VERSION : 0.1
   VAR_INPUT
      OFF_SQ : Bool := false;   // Turn sequence off
      INIT_SQ : Bool := false;   // Set sequence to initial state
      ACK_EF : Bool := false;   // Acknowledge all errors and faults
      S_PREV : Bool := false;   // Output previous step in parameter S_NO
      S_NEXT : Bool := false;   // Indicate next step in parameter S_NO
      SW_AUTO : Bool := false;   // Automatic mode
      SW_TAP : Bool := false;   // Semiautomatic/switch with transition
      SW_TOP : Bool := false;   // Semiautomatic/ignore transition
      SW_MAN : Bool := false;   // Manual mode
      S_SEL : Int := 0;   // Select step to be output to S_NO
      S_ON : Bool := false;   // Activate step indicated in S_NO
      S_OFF : Bool := false;   // Deactivate step indicated S_NO
      T_PUSH : Bool := false;   // Enable transition to switch in semi automatic mode
      "Confimation Position 1" : Bool;
      "Confirmation Position 2" : Bool;
      "Products more than zero" : Bool;
      "Products zero" : Bool;
      "Timer 1" : Time;
   END_VAR
   VAR_OUTPUT
      S_NO : Int := 0;   // Step number
      S_MORE : Bool := false;   // More steps are available and can be shown in S_NO
      S_ACTIVE : Bool := false;   // Step indicated in S_NO is active
      ERR_FLT : Bool := false;   // Interlock or supervision group error
      AUTO_ON : Bool := false;   // Automatic mode is active
      TAP_ON : Bool := false;   // Semiautomatic mode/step with transition enabled
      TOP_ON : Bool := false;   // Semiautomatic mode/ignore transition enabled
      MAN_ON : Bool := false;   // Manual mode is active
      "Move Position 1" : Bool;
      "Move Position 2" : Bool;
   END_VAR
   VAR
      SWITCH : Array[0..0] of DWord;
      SW_SQTS : Array[0..9] of Byte;
      SW_ADDR : Word := 16#E;
      G7T_0 : GraphTransition;
      G7S_0 : GraphStep;
      PRE_CRIT : Array[0..0] of DWord;
      POST_CRIT : Array[0..0] of DWord;
      TVX : Array[0..6] of Byte;
      TTX : Array[0..6] of Byte;
      TSX : Array[0..2] of Byte;
      S00X : Array[0..2] of Byte;
      SOFFX : Array[0..2] of Byte;
      SONX : Array[0..2] of Byte;
      SAX : Array[0..2] of Byte;
      SERRX : Array[0..10] of Byte;
      SMX : Array[0..10] of Byte;
      S0X : Array[0..10] of Byte;
      S1X : Array[0..10] of Byte;
      S_DISPLAY : Int;   // Internal display of output parameter S_NO
      S_SEL_OLD : Int;   // Previous value in S_SEL
      S_DISPIDX : Byte;   // Index of the step in S_NO
      T_DISPIDX : Byte;   // Index of the transition displayed in T_NO
      MOPEDGE : Struct
         AUTO : Bool := false;
         MAN : Bool := false;
         TAP : Bool := false;
         TOP : Bool := false;
         ACK_S : Bool := false;
         REG_S : Bool := false;
         T_PREV : Bool := false;
         T_NEXT : Bool := false;
         LOCK : Bool := false;
         SUP : Bool := false;
         ACKREQ : Bool := false;
         SSKIP : Bool := false;
         OFF : Bool := false;
         INIT : Bool := false;
         HALT : Bool := false;
         TMS_HALT : Bool := false;
         OPS_ZERO : Bool := false;
         SACT_DISP : Bool := false;
         SEF_DISP : Bool := false;
         SALL_DISP : Bool := false;
         S_PREV : Bool := false;
         S_NEXT : Bool := false;
         S_SELOK : Bool := false;
         S_ON : Bool := false;
         S_OFF : Bool := false;
         T_PUSH : Bool := false;
         REG : Bool := false;
         ACK : Bool := false;
         IL_PERM : Bool := false;
         T_PERM : Bool := false;
         ILP_MAN : Bool := false;
      END_STRUCT;
      MOP : Struct   // Mode
         AUTO : Bool := true;   // Status: automatic mode
         MAN : Bool := false;   // Status: manual mode
         TAP : Bool := false;   // Status: semi automatic/switch with transition
         TOP : Bool := false;   // Status: semi automatic/ignore transition
         ACK_S : Bool := false;   // Request: acknowledge step at parameter S_NO
         REG_S : Bool := false;   // Request: register step indicated in S_NO
         T_PREV : Bool := false;   // Request: output previous valid transition in T_NO
         T_NEXT : Bool := false;   // Request: output next valid transition in T_NO
         LOCK : Bool := true;   // Status: interlocks activated
         SUP : Bool := true;   // Status: supervisions activated
         ACKREQ : Bool := true;   // Status: acknowledgment required
         SSKIP : Bool := false;   // Status: "Skip steps" enabled
         OFF : Bool := false;   // Request: deactivate all steps
         INIT : Bool := true;   // Request: set sequence to initial state
         HALT : Bool := false;   // Status: sequence halted
         TMS_HALT : Bool := false;   // Status: all internal timers held
         OPS_ZERO : Bool := false;   // Status: set all operands processed with N, L, D instructions to 0
         SACT_DISP : Bool := true;   // Status: display active steps only
         SEF_DISP : Bool := false;   // Status: display only steps with errors and disrupted steps
         SALL_DISP : Bool := false;   // Status: display all steps
         S_PREV : Bool := false;   // Request: output previous step to S_NO
         S_NEXT : Bool := false;   // Request: Output next step at S_NO parameter
         S_SELOK : Bool := false;   // Request: output step number from S_SEL to S_NO
         S_ON : Bool := false;   // Request: activate step indicated in S_NO
         S_OFF : Bool := false;   // Request: deactivate step at parameter S_NO
         T_PUSH : Bool := false;   // Request: transition switching enabled
         REG : Bool := false;   // Request: register all interlock and supervision errors
         ACK : Bool := false;   // Request: acknowledge all interlock and supervision errors
         IL_PERM : Bool := false;   // Status: permanent processing of all interlocks
         T_PERM : Bool := false;   // Status: permanent processing of all transitions
         ILP_MAN : Bool := false;   // Status: permanent processing of all interlocks in manual mode
      END_STRUCT;
      TICKS : Struct   // Clock speeds
         DELTA : Time := T#0ms;   // Time difference between cycles
         OLD : Time := T#0ms;   // 10 ms clock counter value in last cycle
         NEW : Time := T#0ms;   // 10 ms clock counter value in this cycle
      END_STRUCT;
      SQ_FLAGS : Struct   // Sequence bit memory
         ERR_FLT : Bool := false;   // Interlock and supervision group error
         ERROR : Bool := false;   // Interlock group error
         FAULT : Bool := false;   // Supervision group error
         RT_FAIL : Bool := false;   // Runtime error
         NO_SNO : Bool := false;   // Requested step number not found
         NF_OFL : Bool := false;   // Overflow: too many ON or OFF requests
         SA_OFL : Bool := false;   // Overflow: too many steps active
         TV_OFL : Bool := false;   // Overflow: too many valid transitions
         MSG_OFL : Bool := false;   // Overflow: not enough system resources for ALARM_S
         NO_SWI : Bool := false;   // Do not switch in this cycle
         CYC_OP : Bool := false;   // Cyclic execution of the sequence after initialization
         AS_MSG : Bool := true;   // Alarms during runtime enabled or disabled by instruction
         AS_SEND : Bool := false;   // Send alarms from WR_USMSG or only enter in diagnostics buffer
         SQ_BUSY : Bool := false;   // Internal edge memory bit for sequence processing
         SA_BUSY : Bool := false;   // Internal edge memory bit for sequence processing
         AS_SIG : Bool := false;   // Edge memory bit for alarms from Alarm_S and Alarm_SQ
      END_STRUCT;
      S_PTR : DWord := 16#6F0;
      S_PTR2 : DWord := 16#0;
      S_PTR3 : DWord := 16#1370;
      S_PTR4 : DWord := 16#1310;
      T_PTR : DWord := 16#12B0;
      C_AR2 : DWord := 16#0;
      M_FBDB : DWord := 16#C0000;
      M_SNO : Word := 16#0;
      M_EVID : Word := 16#0;
      M_EVIL : C_Alarm_s;
      M_EVSV : C_Alarm_s;
      M_EV : DWord := 16#11F0;
      CRIT : Array[0..31] of Bool;
      S_START : Byte := 16#0;
      S_IDX : Byte := 16#0;
      S_INT : Int := 72;
      S_TMP : Byte := 16#0;
      T_START : Byte := 16#0;
      T_IDX : Byte := 16#0;
      T_TMP : Byte := 16#0;
      T_TMP2 : Byte := 16#00;
      TV_POT : Byte := 16#0A;
      RETURN1 : Byte := 16#0;
      RETURN2 : Byte := 16#0;
      SINI : Array[0..2] of Byte;
      LSTT : Array[0..11] of Byte;
      ATAJ : Array[0..11] of Byte;
      ATAB : Array[0..11] of Byte;
      PSTT : Array[0..11] of Byte;
      NSTT : Array[0..11] of Byte;
      ASSJ : Array[0..9] of Byte;
      ASSB : Array[0..9] of Byte;
      PTTS : Array[0..9] of Byte;
      NTTS : Array[0..9] of Byte;
      PRE_CNT : Word := 16#1;
      POST_CNT : Word := 16#1;
      ADR_COND : Word := 16#0;
      MAX_TVAL : Byte := 16#5;
      MAX_SACT : Byte := 16#1;
      MAX_CRIT : Byte := 16#4;
      T_CNT : Byte := 16#B;
      SUP_CNT : Byte := 16#0;
      LOCK_CNT : Byte := 16#0;
      S_CNT : Byte := 16#9;
      SQ_CNT : Byte := 16#1;
      PRS_INPAR : DWord := 16#E000FEC8;
      PRS_OUTPAR : DWord := 16#E000800F;
      GC_FLAGS : Struct
         T_MACH : Byte := 16#EB;
         COND_ED : Byte := 16#E3;
         W_LEVEL : Byte := 16#D5;
         FB_IF : Byte := 16#FA;
         AS_MSG : Word := 16#404;
         SSB : Word := 16#108;
         DILG : Word := 16#362;
         ADDR_T0 : Word := 16#1E;
         CRIT_AVAIL : Bool := false;
         SSKIP_AVAIL : Bool := true;
         SSKIP_ON : Bool := false;
         ACK_REQ : Bool := true;
         SYNC_AVAIL : Bool := true;
         ILP_MAN : Bool := false;
         SWM_LOCKED : Bool := false;
         SAVE_SW : Bool := true;
      END_STRUCT;
      G7_FBMARK : Byte := 16#3C;
      G7_RELEASE : Byte := 16#3C;
      G7_ID2 : Byte := 16#37;
      G7_ID1 : Byte := 16#47;
   END_VAR
   // SW_SQTS[0] := 16#3;
   // SW_SQTS[8] := 16#2;
   // SW_SQTS[9] := 16#2;
   // TVX[0] := 16#1;
   // TTX[0] := 16#1;
   // TSX[0] := 16#1;
   // S00X[0] := 16#1;
   // SOFFX[0] := 16#1;
   // SONX[0] := 16#1;
   // SAX[0] := 16#1;
   // SERRX[0] := 16#1;
   // SMX[0] := 16#1;
   // S0X[0] := 16#1;
   // S1X[0] := 16#1;
   // SINI[0] := 16#2;
   // SINI[1] := 16#1;
   // SINI[2] := 0;
   // LSTT[0] := 0;
   // LSTT[1] := 0;
   // LSTT[2] := 0;
   // LSTT[3] := 0;
   // LSTT[4] := 0;
   // LSTT[5] := 0;
   // LSTT[6] := 0;
   // LSTT[7] := 16#4;
   // LSTT[8] := 0;
   // LSTT[9] := 0;
   // LSTT[10] := 16#1;
   // ATAJ[0] := 0;
   // ATAJ[1] := 16#1;
   // ATAJ[2] := 16#2;
   // ATAJ[3] := 16#3;
   // ATAJ[4] := 16#4;
   // ATAJ[5] := 16#5;
   // ATAJ[6] := 16#6;
   // ATAJ[7] := 16#7;
   // ATAJ[8] := 16#8;
   // ATAJ[9] := 16#9;
   // ATAJ[10] := 16#A;
   // ATAB[0] := 0;
   // ATAB[1] := 16#1;
   // ATAB[2] := 16#2;
   // ATAB[3] := 16#B;
   // ATAB[4] := 16#4;
   // ATAB[5] := 16#5;
   // ATAB[6] := 16#6;
   // ATAB[7] := 16#8;
   // ATAB[8] := 16#7;
   // ATAB[9] := 16#9;
   // ATAB[10] := 16#A;
   // PSTT[0] := 0;
   // PSTT[1] := 16#1;
   // PSTT[2] := 16#2;
   // PSTT[3] := 16#3;
   // PSTT[4] := 16#4;
   // PSTT[5] := 16#5;
   // PSTT[6] := 16#6;
   // PSTT[7] := 16#7;
   // PSTT[8] := 16#7;
   // PSTT[9] := 16#8;
   // PSTT[10] := 16#9;
   // NSTT[0] := 16#1;
   // NSTT[1] := 16#2;
   // NSTT[2] := 16#3;
   // NSTT[3] := 16#4;
   // NSTT[4] := 16#5;
   // NSTT[5] := 16#6;
   // NSTT[6] := 16#7;
   // NSTT[7] := 16#4;
   // NSTT[8] := 16#8;
   // NSTT[9] := 16#9;
   // NSTT[10] := 16#1;
   // ASSJ[0] := 0;
   // ASSJ[1] := 16#1;
   // ASSJ[2] := 16#2;
   // ASSJ[3] := 16#3;
   // ASSJ[4] := 16#4;
   // ASSJ[5] := 16#5;
   // ASSJ[6] := 16#6;
   // ASSJ[7] := 16#7;
   // ASSJ[8] := 16#8;
   // ASSJ[9] := 16#9;
   // ASSB[0] := 0;
   // ASSB[1] := 16#1;
   // ASSB[2] := 16#2;
   // ASSB[3] := 16#3;
   // ASSB[4] := 16#4;
   // ASSB[5] := 16#5;
   // ASSB[6] := 16#6;
   // ASSB[7] := 16#7;
   // ASSB[8] := 16#8;
   // ASSB[9] := 16#9;
   // PTTS[0] := 0;
   // PTTS[2] := 16#1;
   // PTTS[3] := 16#2;
   // PTTS[4] := 16#3;
   // PTTS[5] := 16#4;
   // PTTS[6] := 16#5;
   // PTTS[7] := 16#6;
   // PTTS[8] := 16#8;
   // PTTS[9] := 16#9;
   // NTTS[0] := 0;
   // NTTS[1] := 16#1;
   // NTTS[2] := 16#2;
   // NTTS[3] := 16#3;
   // NTTS[4] := 16#4;
   // NTTS[5] := 16#5;
   // NTTS[6] := 16#6;
   // NTTS[7] := 16#7;
   // NTTS[8] := 16#9;
   // NTTS[9] := 16#A;
   // SW_SQTS[4] := 16#1;
   // SW_SQTS[5] := 16#1;
   // SW_SQTS[6] := 16#1;
   // SW_SQTS[7] := 16#1;
   // LSTT[11] := 16#1;
   // ATAJ[11] := 16#B;
   // ATAB[11] := 16#3;
   // PSTT[11] := 16#3;
   // NSTT[11] := 16#1;
BEGIN
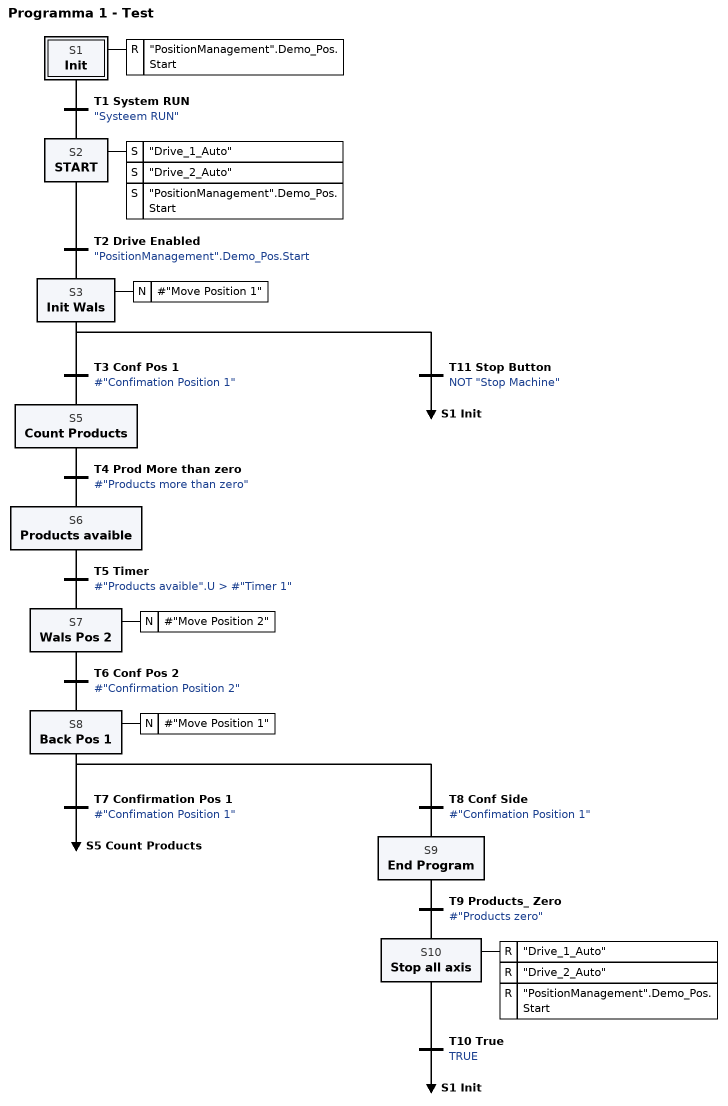
   // sequencer 1
   INITIAL_STEP Init:   // S1
              R    "PositionManagement".Demo_Pos.Start
   END_STEP
   TRANSITION "System RUN" FROM Init TO START   // T1
      := "Systeem RUN";
   END_TRANSITION
   STEP START:   // S2
      // Set Ouputs
              S    "Drive_1_Auto"
              S    "Drive_2_Auto"
              S    "PositionManagement".Demo_Pos.Start
   END_STEP
   TRANSITION "Drive Enabled" FROM START TO "Init Wals"   // T2
      := "PositionManagement".Demo_Pos.Start;
   END_TRANSITION
   STEP "Init Wals":   // S3
      // Move Start Position4
              N    #"Move Position 1"
   END_STEP
   TRANSITION "Conf Pos 1" FROM "Init Wals" TO "Count Products"   // T3
      := #"Confimation Position 1";
   END_TRANSITION
   TRANSITION "Stop Button" FROM "Init Wals" TO Init   // T11, jump
      := NOT "Stop Machine";
   END_TRANSITION
   STEP "Count Products":   // S5
   END_STEP
   TRANSITION "Prod More than zero" FROM "Count Products" TO "Products avaible"   // T4
      := #"Products more than zero";
   END_TRANSITION
   STEP "Products avaible":   // S6
   END_STEP
   TRANSITION "Timer" FROM "Products avaible" TO "Wals Pos 2"   // T5: Timer 1
      := #"Products avaible".U > #"Timer 1";
   END_TRANSITION
   STEP "Wals Pos 2":   // S7
              N    #"Move Position 2"
   END_STEP
   TRANSITION "Conf Pos 2" FROM "Wals Pos 2" TO "Back Pos 1"   // T6
      := #"Confirmation Position 2";
   END_TRANSITION
   STEP "Back Pos 1":   // S8
      // Move Position 1
              N    #"Move Position 1"
   END_STEP
   TRANSITION "Confirmation Pos 1" FROM "Back Pos 1" TO "Count Products"   // T7, jump: Conf Pos 1
      := #"Confimation Position 1";
   END_TRANSITION
   TRANSITION "Conf Side" FROM "Back Pos 1" TO "End Program"   // T8
      := #"Confimation Position 1";
   END_TRANSITION
   STEP "End Program":   // S9
   END_STEP
   TRANSITION "Products_ Zero" FROM "End Program" TO "Stop all axis"   // T9
      := #"Products zero";
   END_TRANSITION
   STEP "Stop all axis":   // S10
      // Reset Axis
              R    "Drive_1_Auto"
              R    "Drive_2_Auto"
              R    "PositionManagement".Demo_Pos.Start
   END_STEP
   TRANSITION True FROM "Stop all axis" TO Init   // T10, jump
      := TRUE;
   END_TRANSITION
END_FUNCTION_BLOCK

FUNCTION_BLOCK "FB_ProductTrigger"   // FB13, SCL
{ S7_Optimized_Access := 'FALSE' }
VERSION : 0.1
   VAR_INPUT
      SensorInput : Bool;
      TimeDelay : Time;
      SystemTime : Time;
   END_VAR
   VAR_OUTPUT
      TriggerMovement : Bool;
      ProductCount : Int;
   END_VAR
   VAR_TEMP
      ProductQueue : Array[0..1] of "ProductEntry";
      SensorMemory : Bool;
      i : Int;
   END_VAR
BEGIN
   // Reset output
   #TriggerMovement := FALSE;

   // Flankdetectie op sensor
   IF #SensorInput AND NOT #SensorMemory THEN
       // Zoek eerste vrije plek
       FOR #i := 1 TO 10 DO
           IF NOT #ProductQueue[#i].Active THEN
               #ProductQueue[#i].Active := TRUE;
               #ProductQueue[#i].StartTime := #SystemTime;
               EXIT;
           END_IF;
       END_FOR;
   END_IF;
   #SensorMemory := #SensorInput;

   // Kijk of een van de producten klaar is voor beweging
   FOR #i := 1 TO 10 DO
       IF #ProductQueue[#i].Active AND (#SystemTime - #ProductQueue[#i].StartTime >= #TimeDelay) THEN
           #TriggerMovement := TRUE;
           #ProductQueue[#i].Active := FALSE; // Verwijder uit wachtrij
           EXIT; // Eén tegelijk
       END_IF;
   END_FOR;

   // Update productenteller
   #ProductCount := 0;
   FOR #i := 1 TO 10 DO
       IF #ProductQueue[#i].Active THEN
           #ProductCount := #ProductCount + 1;
       END_IF;
   END_FOR;
END_FUNCTION_BLOCK

FUNCTION_BLOCK "FB_SystemTimeCounter"   // FB14, SCL
{ S7_Optimized_Access := 'FALSE' }
VERSION : 0.1
   VAR_INPUT
      Enable : Bool;
      CycleTime : Time;
   END_VAR
   VAR_OUTPUT
      SystemTime : Time;
   END_VAR
   VAR_TEMP
      PrevEnable : Bool;
   END_VAR
BEGIN
   //Start//

   IF #Enable THEN
       // Enkel verhogen als Enable TRUE is
       #SystemTime := #SystemTime + #CycleTime;
   END_IF;

   // Reset eventueel bij FALSE->TRUE flank
   //IF NOT #PrevEnable AND #Enable THEN
       // Optioneel reset: SystemTime := T#0s;
   //END_IF;

   #PrevEnable := #Enable;
END_FUNCTION_BLOCK

FUNCTION_BLOCK "Blinker"   // FB15, SCL
{ S7_Optimized_Access := 'FALSE' }
VERSION : 0.1
   VAR_INPUT
      Enable : Bool;
      BlinkTime : Time := T#500ms;
   END_VAR
   VAR_OUTPUT
      Q_Blink : Bool;
      Q_Blink2 : Bool;
   END_VAR
   VAR
      BlinkTimer : TON;
   END_VAR
   VAR_TEMP
      LastToggleTime : Time;
   END_VAR
BEGIN
   // Logica
   IF #Enable THEN
       #BlinkTimer(IN := TRUE,
                   PT := #BlinkTime);   // Correct gebruik van PT

       IF #BlinkTimer.Q THEN
           #Q_Blink := NOT #Q_Blink;                // Toggle uitgang
           #Q_Blink2 := NOT #Q_Blink2;
           #BlinkTimer(IN := FALSE,
                       PT := #BlinkTime); // Reset timer (verplicht opnieuw PT meegeven)
       END_IF;

   ELSE
       #BlinkTimer(IN := FALSE,
                   PT := #BlinkTime);  // Timer uitzetten
       #Q_Blink := FALSE; // Uitgang terug laag
       #Q_Blink2 := FALSE;
   END_IF;
END_FUNCTION_BLOCK

FUNCTION_BLOCK "BlowOff_Timer"   // FB16, SCL
{ S7_Optimized_Access := 'FALSE' }
VERSION : 0.1
   VAR_INPUT
      Enable : Bool;
      CycleTime : Time;
      PulseDuration : Time;
      NowTime : Time;
   END_VAR
   VAR_OUTPUT
      Q_Pulse : Bool;
   END_VAR
   VAR
      CycleTimer : TON;
      PulseTimer : TON;
      State : Int;
      S_PEXT : Int;
   END_VAR
   VAR_TEMP
      PulseActive : Bool;
      StartPulse : Bool;
      TriggerPulse : Bool;
      PulseBusy : Bool;
      DummyWord : Word;
      DummyWord2 : Bool;
      T1 : Int;
      PulseStartTime : Time;
      LastPulseEndTime : Time;
      LastPulseTime : Time;
   END_VAR
BEGIN
   // Logica
   IF #Enable THEN
       // Start cyclische timer
       #CycleTimer(IN := TRUE,
                   PT := #CycleTime);

       IF #CycleTimer.Q THEN
           // Start puls-timer als cyclus voorbij is
           #PulseTimer(IN := TRUE,
                       PT := #PulseDuration);

           // Reset de CycleTimer voor de volgende cyclus
           #CycleTimer(IN := FALSE,
                       PT := #CycleTime);
       END_IF;

       // Puls-timer logica
       IF #PulseTimer.IN THEN
           #Q_Pulse := TRUE;

           IF #PulseTimer.Q THEN
               // Puls voorbij, pulse output uit
               #PulseTimer(IN := FALSE,
                           PT := #PulseDuration);
               #Q_Pulse := FALSE;
           END_IF;
       ELSE
           #Q_Pulse := FALSE;
       END_IF;

   ELSE
       // Alles resetten bij disable
       #CycleTimer(IN := FALSE,
                   PT := #CycleTime);
       #PulseTimer(IN := FALSE,
                   PT := #PulseDuration);
       #Q_Pulse := FALSE;
   END_IF;
END_FUNCTION_BLOCK

FUNCTION_BLOCK "ProductBuffer"   // FB17, SCL
{ S7_Optimized_Access := 'FALSE' }
VERSION : 0.1
   VAR_INPUT
      SensorInput : Bool;
      TimeDelay : Time;
      TriggerFeedback : Bool;
   END_VAR
   VAR_OUTPUT
      TriggerMovement : Bool;
      ProductCount : Int;
   END_VAR
   VAR
      PrevSensor : Bool;
      DelayTimer : TON;
      MovementActive : Bool;
   END_VAR
BEGIN
   // Flankdetectie op sensor
   IF #SensorInput AND NOT #PrevSensor THEN
       IF #ProductCount < 32767 THEN
           #ProductCount := #ProductCount + 1;
       END_IF;
   END_IF;
   #PrevSensor := #SensorInput;

   // Timer mag alleen lopen als:
   // - Er producten zijn
   // - Er geen beweging actief is
   IF (#ProductCount > 0) AND (NOT #MovementActive) THEN
       #DelayTimer(IN := TRUE,
                   PT := #TimeDelay);
   ELSE
       #DelayTimer(IN := FALSE,
                   PT := #TimeDelay);
   END_IF;

   // Als de timer klaar is → activeer beweging en zet MovementActive
   IF #DelayTimer.Q THEN
       #TriggerMovement := TRUE;
       #MovementActive := TRUE;
       #ProductCount := #ProductCount - 1;
       #DelayTimer(IN := FALSE,
                   PT := #TimeDelay); // Reset timer
   END_IF;

   // Wacht op TriggerFeedback om TriggerMovement terug laag te zetten
   IF #MovementActive AND #TriggerFeedback THEN
       #TriggerMovement := FALSE;
       #MovementActive := FALSE;
   END_IF;
END_FUNCTION_BLOCK

FUNCTION_BLOCK "ProductBuffer_V2"   // FB18, SCL
{ S7_Optimized_Access := 'FALSE' }
VERSION : 0.1
   VAR_INPUT
      SensorInput : Bool;
      SensorManual : Bool;
      TimeDelay : Time;
      SystemTime : Time;
      TriggerFeedback : Bool;
   END_VAR
   VAR_OUTPUT
      TriggerMovement : Bool;
      InsertIndex : Int;
      ProductCount : Int;
      SystemTicks : DInt;
   END_VAR
   VAR
      ProductQueue : Array[0..1] of "ProductEntry";
      StartTimes : Struct
         _0 : Time;
         _1 : Time;
         _2 : Time;
         _3 : Time;
         _4 : Time;
         _5 : Time;
         _6 : Time;
         _7 : Time;
         _8 : Time;
         _9 : Time;
      END_STRUCT;
      Actives : Struct
         _0 : Bool;
         _1 : Bool;
         _2 : Bool;
         _3 : Bool;
         _4 : Bool;
         _5 : Bool;
         _6 : Bool;
         _7 : Bool;
         _8 : Bool;
         _9 : Bool;
      END_STRUCT;
      PrevSensor : Bool;
      MovementActive : Bool;
      i : Int;
      Elapsed : DInt;
   END_VAR
BEGIN
   // Flankdetectie sensor
   IF #SensorInput AND NOT #PrevSensor THEN
       CASE #InsertIndex MOD 10 OF
           0:
               IF NOT #Actives._0 THEN
                   #Actives._0 := TRUE;
                   #StartTimes._0 := #SystemTime;
               END_IF;
           1:
               IF NOT #Actives._1 THEN
                   #Actives._1 := TRUE;
                   #StartTimes._1 := #SystemTime;
               END_IF;
           2:
               IF NOT #Actives._2 THEN
                   #Actives._2 := TRUE;
                   #StartTimes._2 := #SystemTime;
               END_IF;
           3:
               IF NOT #Actives._3 THEN
                   #Actives._3 := TRUE;
                   #StartTimes._3 := #SystemTime;
               END_IF;
           4:
               IF NOT #Actives._4 THEN
                   #Actives._4 := TRUE;
                   #StartTimes._4 := #SystemTime;
               END_IF;
           5:
               IF NOT #Actives._5 THEN
                   #Actives._5 := TRUE;
                   #StartTimes._5 := #SystemTime;
               END_IF;
           6:
               IF NOT #Actives._6 THEN
                   #Actives._6 := TRUE;
                   #StartTimes._6 := #SystemTime;
               END_IF;
           7:
               IF NOT #Actives._7 THEN
                   #Actives._7 := TRUE;
                   #StartTimes._7 := #SystemTime;
               END_IF;
           8:
               IF NOT #Actives._8 THEN
                   #Actives._8 := TRUE;
                   #StartTimes._8 := #SystemTime;
               END_IF;
           9:
               IF NOT #Actives._9 THEN
                   #Actives._9 := TRUE;
                   #StartTimes._9 := #SystemTime;
               END_IF;
       END_CASE;
       #InsertIndex := (#InsertIndex + 1) MOD 10;
   END_IF;

   #PrevSensor := #SensorInput;

   // Tellen hoeveel producten actief zijn
   #ProductCount := 0;
   IF #Actives._0 THEN
       #ProductCount := #ProductCount + 1;
   END_IF;
   IF #Actives._1 THEN
       #ProductCount := #ProductCount + 1;
   END_IF;
   IF #Actives._2 THEN
       #ProductCount := #ProductCount + 1;
   END_IF;
   IF #Actives._3 THEN
       #ProductCount := #ProductCount + 1;
   END_IF;
   IF #Actives._4 THEN
       #ProductCount := #ProductCount + 1;
   END_IF;
   IF #Actives._5 THEN
       #ProductCount := #ProductCount + 1;
   END_IF;
   IF #Actives._6 THEN
       #ProductCount := #ProductCount + 1;
   END_IF;
   IF #Actives._7 THEN
       #ProductCount := #ProductCount + 1;
   END_IF;
   IF #Actives._8 THEN
       #ProductCount := #ProductCount + 1;
   END_IF;
   IF #Actives._9 THEN
       #ProductCount := #ProductCount + 1;
   END_IF;

   // Beweging starten als een product klaar is en geen andere beweging actief is
   IF NOT #MovementActive THEN
       IF #Actives._0 THEN
           #Elapsed := TIME_TO_DINT(#SystemTime) - TIME_TO_DINT(#StartTimes._0);
           IF #Elapsed >= TIME_TO_DINT(#TimeDelay) THEN
               #TriggerMovement := TRUE;
               #MovementActive := TRUE;
               #Actives._0 := FALSE;
           END_IF;
       ELSIF #Actives._1 THEN
           #Elapsed := TIME_TO_DINT(#SystemTime) - TIME_TO_DINT(#StartTimes._1);
           IF #Elapsed >= TIME_TO_DINT(#TimeDelay) THEN
               #TriggerMovement := TRUE;
               #MovementActive := TRUE;
               #Actives._1 := FALSE;
           END_IF;
       ELSIF #Actives._2 THEN
           #Elapsed := TIME_TO_DINT(#SystemTime) - TIME_TO_DINT(#StartTimes._2);
           IF #Elapsed >= TIME_TO_DINT(#TimeDelay) THEN
               #TriggerMovement := TRUE;
               #MovementActive := TRUE;
               #Actives._2 := FALSE;
           END_IF;
       ELSIF #Actives._3 THEN
           #Elapsed := TIME_TO_DINT(#SystemTime) - TIME_TO_DINT(#StartTimes._3);
           IF #Elapsed >= TIME_TO_DINT(#TimeDelay) THEN
               #TriggerMovement := TRUE;
               #MovementActive := TRUE;
               #Actives._3 := FALSE;
           END_IF;
       ELSIF #Actives._4 THEN
           #Elapsed := TIME_TO_DINT(#SystemTime) - TIME_TO_DINT(#StartTimes._4);
           IF #Elapsed >= TIME_TO_DINT(#TimeDelay) THEN
               #TriggerMovement := TRUE;
               #MovementActive := TRUE;
               #Actives._4 := FALSE;
           END_IF;
       ELSIF #Actives._5 THEN
           #Elapsed := TIME_TO_DINT(#SystemTime) - TIME_TO_DINT(#StartTimes._5);
           IF #Elapsed >= TIME_TO_DINT(#TimeDelay) THEN
               #TriggerMovement := TRUE;
               #MovementActive := TRUE;
               #Actives._5 := FALSE;
           END_IF;
       ELSIF #Actives._6 THEN
           #Elapsed := TIME_TO_DINT(#SystemTime) - TIME_TO_DINT(#StartTimes._6);
           IF #Elapsed >= TIME_TO_DINT(#TimeDelay) THEN
               #TriggerMovement := TRUE;
               #MovementActive := TRUE;
               #Actives._6 := FALSE;
           END_IF;
       ELSIF #Actives._7 THEN
           #Elapsed := TIME_TO_DINT(#SystemTime) - TIME_TO_DINT(#StartTimes._7);
           IF #Elapsed >= TIME_TO_DINT(#TimeDelay) THEN
               #TriggerMovement := TRUE;
               #MovementActive := TRUE;
               #Actives._7 := FALSE;
           END_IF;
       ELSIF #Actives._8 THEN
           #Elapsed := TIME_TO_DINT(#SystemTime) - TIME_TO_DINT(#StartTimes._8);
           IF #Elapsed >= TIME_TO_DINT(#TimeDelay) THEN
               #TriggerMovement := TRUE;
               #MovementActive := TRUE;
               #Actives._8 := FALSE;
           END_IF;
       ELSIF #Actives._9 THEN
           #Elapsed := TIME_TO_DINT(#SystemTime) - TIME_TO_DINT(#StartTimes._9);
           IF #Elapsed >= TIME_TO_DINT(#TimeDelay) THEN
               #TriggerMovement := TRUE;
               #MovementActive := TRUE;
               #Actives._9 := FALSE;
           END_IF;
       END_IF;
   END_IF;

   // Beweging beëindigen na feedback
   IF #MovementActive AND #TriggerFeedback THEN
       #TriggerMovement := FALSE;
       #MovementActive := FALSE;
   END_IF;
END_FUNCTION_BLOCK

FUNCTION_BLOCK "ProductBuffer_V3"   // FB20, SCL
{ S7_Optimized_Access := 'FALSE' }
VERSION : 0.1
   VAR_INPUT
      SensorInput : Bool;   // Sensor aan begin band
      EncoderPosition : Real;   // Koppel aan Encoder Data Instance
      TriggerDistance : Real;   // Gewenste Afstand Product voor trigger
      TriggerFeedback : Bool;
   END_VAR
   VAR_OUTPUT
      TriggerMovement : Bool;   // Trigger Start Movement
      ProductCount : Int;   // Count products in buffer
   END_VAR
   VAR
      ProductBuffer : Array[0..9] of "ProductTrack";
      PrevSensor : Bool;
      MovementActive : Bool;
      i : Int;
      Distance : Real;
   END_VAR
BEGIN
   // 1️⃣ Flankdetectie - detecteer nieuw product
   IF #SensorInput AND NOT #PrevSensor THEN
       FOR #i := 0 TO 9 DO
           IF NOT #ProductBuffer[#i].Active THEN
               #ProductBuffer[#i].StartPosition := #EncoderPosition;
               #ProductBuffer[#i].Active := TRUE;
               EXIT;
           END_IF;
       END_FOR;
   END_IF;
   #PrevSensor := #SensorInput;

   // 2️⃣ Tel actieve producten
   #ProductCount := 0;
   FOR #i := 0 TO 9 DO
       IF #ProductBuffer[#i].Active THEN
           #ProductCount := #ProductCount + 1;
       END_IF;
   END_FOR;

   // 3️⃣ Zoek eerste product dat zijn afstand heeft afgelegd
   IF NOT #MovementActive THEN
       FOR #i := 0 TO 9 DO
           IF #ProductBuffer[#i].Active THEN
               #Distance := #EncoderPosition - #ProductBuffer[#i].StartPosition;

               IF #Distance >= #TriggerDistance THEN
                   #TriggerMovement := TRUE;
                   #MovementActive := TRUE;
                   #ProductBuffer[#i].Active := FALSE;
                   EXIT;
               END_IF;
           END_IF;
       END_FOR;
   END_IF;

   // 4️⃣ Wacht op feedback om beweging af te ronden
   IF #MovementActive AND #TriggerFeedback THEN
       #TriggerMovement := FALSE;
       #MovementActive := FALSE;
   END_IF;
END_FUNCTION_BLOCK

FUNCTION "SCL_Block" : Void   // FC10, SCL
{ S7_Optimized_Access := 'FALSE' }
VERSION : 0.1
BEGIN
   // Reset de Word variabelen aan het begin van elke cyclus
   "Alarms".AlarmsWord := 0;
   "Alarms".HMI_Alarm_Drive1 := 0;
   "Alarms".HMI_Alarm_Drive2 := 0;
   "Alarms".HMI_Alarm_Drive3 := 0;
   "Alarms".HMI_Alarm_Drive4 := 0;
   "Alarms".HMI_Alarm_Drive5 := 0;

   // Controleer de alarmen en zet de respectievelijke bits aan
   IF "Alarms".AlarmStruct.Alarm_Product_Not_Position THEN
       "Alarms".AlarmsWord := "Alarms".AlarmsWord OR WORD#1; // Zet bit 0 aan
   END_IF;

   IF "Alarms".AlarmStruct.Alarm_Axis_Not_Position THEN
       "Alarms".AlarmsWord := "Alarms".AlarmsWord OR WORD#2; // Zet bit 1 aan
   END_IF;

   IF "Alarms".AlarmStruct.Alarm_Drive1 THEN
       "Alarms".HMI_Alarm_Drive1 := "Alarms".HMI_Alarm_Drive1 OR WORD#1; // Zet bit 2 aan
   END_IF;

   IF "Alarms".AlarmStruct.Alarm_Drive2 THEN
       "Alarms".HMI_Alarm_Drive2 := "Alarms".HMI_Alarm_Drive2 OR WORD#1; // Zet bit 3 aan
   END_IF;

   IF "Alarms".AlarmStruct.Alarm_Drive3 THEN
       "Alarms".HMI_Alarm_Drive3 := "Alarms".HMI_Alarm_Drive3 OR WORD#1; // Zet bit 4 aan
   END_IF;

   IF "Alarms".AlarmStruct.Alarm_Drive4 THEN
       "Alarms".HMI_Alarm_Drive4 := "Alarms".HMI_Alarm_Drive4 OR WORD#1; // Zet bit 5 aan
   END_IF;

   IF "Alarms".AlarmStruct.Alarm_Drive5 THEN
       "Alarms".HMI_Alarm_Drive5 := "Alarms".HMI_Alarm_Drive5 OR WORD#1; // Zet bit 6 aan
   END_IF;


   // Position Program Axis 3 (Wals)

   // Configureer de timer om elke 0,5 seconde af te lopen
   "Timer_0_5s".TON(IN := TRUE,
   PT := "PLCMemory"."Encoder PulsOffset");

   // Controleer of de timer is afgelopen
   IF "Timer_0_5s".Q THEN
       // Verhoog of verlaag de positie afhankelijk van de aandrijfsignalen
       IF "Drive 3 RUN FWD" THEN
           "PLCMemory".EncoderPosition := "PLCMemory".EncoderPosition + "PLCMemory".StepSize; // Verhoog met de stepgrootte
       ELSIF "Drive 3 REV" THEN
           "PLCMemory".EncoderPosition := "PLCMemory".EncoderPosition - "PLCMemory".StepSize; // Verlaag met de stepgrootte
       END_IF;

       // Wrapping van de positie bij overschrijden van 360 graden of onder 0 graden
       IF "PLCMemory".EncoderPosition >= 360.0 THEN
           "PLCMemory".EncoderPosition := 0.0;  // Wrapping naar 0 als de positie 360 overschrijdt
       ELSIF "PLCMemory".EncoderPosition < 0.0 THEN
           "PLCMemory".EncoderPosition := 360.0; // Wrapping naar 360 als de positie onder 0 gaat
       END_IF;

       // Reset de timer
       "Timer_0_5s".TON (IN := FALSE,
                         PT := "PLCMemory"."Encoder PulsOffset"); // Reset de timer zodat deze opnieuw kan starten
   END_IF;

   // Homing logica
   IF "Sensor Wals (Option)" THEN
       "PLCMemory".EncoderPosition := 0.0;  // Reset de positie naar 0 als de sensor wordt geactiveerd
   END_IF;



   //Drive Servo Control Here:
   /// Desired Position Axis 3

   // Controleer of de HMI-knop is ingedrukt en er een gewenste positie is ingesteld
   //IF "HMI_Des_Pos_Axis3" THEN
       //"GoButtonPressed" := TRUE; // HMI-knop is ingedrukt, start beweging
   //END_IF;

   // Beveiliging voor de Desired_Encoder_Position: Zorg dat de waarde tussen 0 en 360 blijft
   //IF "PLCMemory".Desired_Encoder_Position > 360.0 THEN
     //  "PLCMemory".Desired_Encoder_Position := 360.0;  // Zet naar 360 als de waarde boven 360 ligt
   //ELSIF "PLCMemory".Desired_Encoder_Position < 0.0 THEN
       //"PLCMemory".Desired_Encoder_Position := 0.0;  // Zet naar 0 als de waarde onder 0 ligt
   //END_IF;

   // Wrapping van de gewenste positie: Als de gewenste positie 360 is, zet deze dan op 0
   //IF "PLCMemory".Desired_Encoder_Position = 360.0 THEN
      // "PLCMemory".Desired_Encoder_Position := 0.0;  // Wrapping naar 0 als de gewenste positie 360 is
   //END_IF;

   // Voer beweging uit totdat de gewenste positie is bereikt
   //IF "GoButtonPressed" THEN
       // Bepaal de bewegingsrichting en start de beweging
     //  IF "PLCMemory".EncoderPosition < "PLCMemory".Desired_Encoder_Position - "PLCMemory".Tolerance THEN
           // Beweeg vooruit met StepSize als snelheid
         //  "PLCMemory".EncoderPosition := "PLCMemory".EncoderPosition + "PLCMemory".StepSize;
        //   "Drive_3_Manual" := TRUE;   // Activeer vooruitbeweging
         //  "Drive 3 REV" := FALSE;     // Zorg dat achteruitbeweging uit is

     //  ELSIF "PLCMemory".EncoderPosition > "PLCMemory".Desired_Encoder_Position + "PLCMemory".Tolerance THEN
           // Beweeg achteruit met StepSize als snelheid
        //   "PLCMemory".EncoderPosition := "PLCMemory".EncoderPosition - "PLCMemory".StepSize;
       //    "Drive_3_Manual" := FALSE;  // Zorg dat vooruitbeweging uit is
       //    "Drive 3 REV" := TRUE;      // Activeer achteruitbeweging

      // ELSE
           // Stop de beweging zodra de positie binnen de tolerantie komt
         //  "Drive_3_Manual" := FALSE;    // Zet vooruitbeweging uit
        //   "Drive 3 REV" := FALSE;       // Zet achteruitbeweging uit
        //   "GoButtonPressed" := FALSE;   // Zet de Go-knop uit om verdere beweging te stoppen
      // END_IF;
   //END_IF;
END_FUNCTION

FUNCTION "SafetyFunction_Block" : Void   // FC12, LAD
{ S7_Optimized_Access := 'FALSE' }
VERSION : 0.1
   VAR_INPUT
      "ESB NC Contact" : Bool;
      "ESB NO Contact" : Bool;
      "Reset NO Contact" : Bool;
      "SAFE door 1 NC Contact" : Bool;
      "SAFE door 2 NC Contact" : Bool;
      "Safety Relais NO Contact" : Bool;
   END_VAR
   VAR_OUTPUT
      SAFE_OK_Signal : Bool;
   END_VAR
BEGIN

REGION Network 1: +MC-21K6:1 - Noodstop Circuit
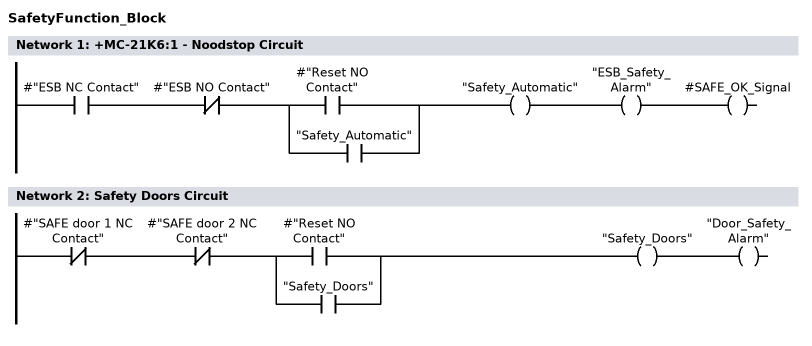
   RUNG wire#powerrail
      Contact( #"ESB NC Contact" )
      I_Contact( #"ESB NO Contact" )
      wire#w1
      Contact( #"Reset NO Contact" )
      wire#w2
      Coil( "Safety_Automatic" )
      Coil( "ESB_Safety_Alarm" )
      Coil( #SAFE_OK_Signal )
   END_RUNG
   RUNG wire#w1
      Contact( "Safety_Automatic" )
   END_RUNG wire#w2
   // the same network as SCL:
   "Safety_Automatic" := #"ESB NC Contact" AND NOT #"ESB NO Contact" AND (#"Reset NO Contact" OR "Safety_Automatic");
   "ESB_Safety_Alarm" := "Safety_Automatic";
   #SAFE_OK_Signal := "Safety_Automatic";
END_REGION

REGION Network 2: Safety Doors Circuit
   RUNG wire#powerrail
      I_Contact( #"SAFE door 1 NC Contact" )
      I_Contact( #"SAFE door 2 NC Contact" )
      wire#w1
      Contact( #"Reset NO Contact" )
      wire#w2
      Coil( "Safety_Doors" )
      Coil( "Door_Safety_Alarm" )
   END_RUNG
   RUNG wire#w1
      Contact( "Safety_Doors" )
   END_RUNG wire#w2
   // the same network as SCL:
   "Safety_Doors" := NOT #"SAFE door 1 NC Contact" AND NOT #"SAFE door 2 NC Contact" AND (#"Reset NO Contact" OR "Safety_Doors");
   "Door_Safety_Alarm" := "Safety_Doors";
END_REGION
END_FUNCTION

FUNCTION "SystemRUN_Block" : Void   // FC13, LAD
{ S7_Optimized_Access := 'FALSE' }
VERSION : 0.1
   VAR_INPUT
      "Safety Relais Contact" : Bool;
      "Stop Machine NC Contact" : Bool;
      "Fill Magzine Contact" : Bool;
      "Start Machine NO Contact" : Bool;
   END_VAR
   VAR_OUTPUT
      "Run Output Lamp" : Bool;
   END_VAR
BEGIN

REGION Network 1: Systeem RUN
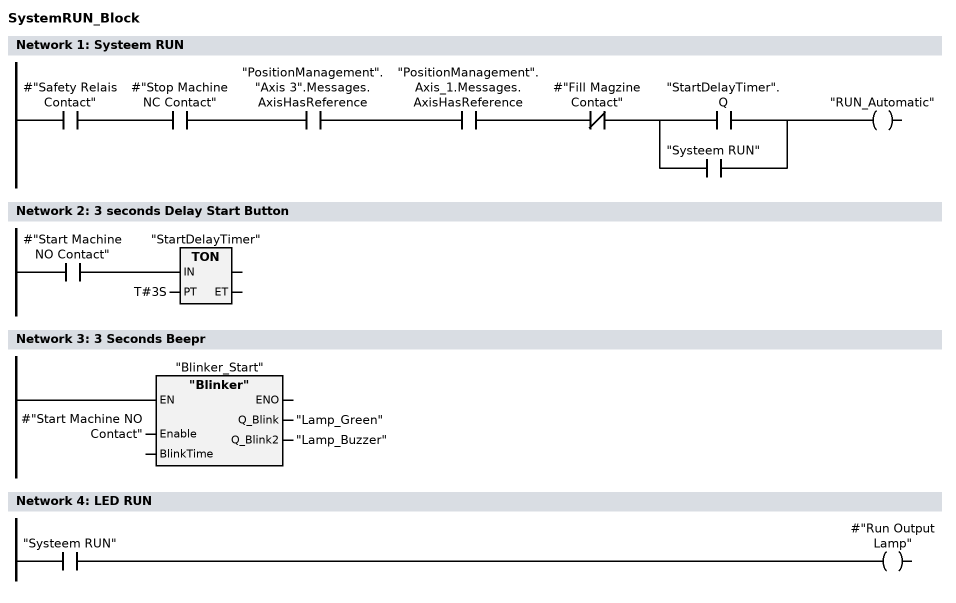
   RUNG wire#powerrail
      Contact( #"Safety Relais Contact" )
      Contact( #"Stop Machine NC Contact" )
      Contact( "PositionManagement"."Axis 3".Messages.AxisHasReference )
      Contact( "PositionManagement".Axis_1.Messages.AxisHasReference )
      I_Contact( #"Fill Magzine Contact" )
      wire#w1
      Contact( "StartDelayTimer".Q )
      wire#w2
      Coil( "RUN_Automatic" )
   END_RUNG
   RUNG wire#w1
      Contact( "Systeem RUN" )
   END_RUNG wire#w2
   // the same network as SCL:
   "RUN_Automatic" := #"Safety Relais Contact" AND #"Stop Machine NC Contact" AND "PositionManagement"."Axis 3".Messages.AxisHasReference AND "PositionManagement".Axis_1.Messages.AxisHasReference AND NOT #"Fill Magzine Contact" AND ("StartDelayTimer".Q OR "Systeem RUN");
END_REGION

REGION Network 2: 3 seconds Delay Start Button
   "StartDelayTimer".TON(IN := #"Start Machine NO Contact", PT := T#3S);
END_REGION

REGION Network 3: 3 Seconds Beepr
   RUNG wire#powerrail
      "Blinker_Start"(Enable := #"Start Machine NO Contact", BlinkTime :=, Q_Blink => "Lamp_Green", Q_Blink2 => "Lamp_Buzzer")
   END_RUNG
   // the same network as SCL:
   "Blinker_Start"(Enable := #"Start Machine NO Contact", Q_Blink => "Lamp_Green", Q_Blink2 => "Lamp_Buzzer");   // "Blinker"
END_REGION

REGION Network 4: LED RUN
   RUNG wire#powerrail
      Contact( "Systeem RUN" )
      Coil( #"Run Output Lamp" )
   END_RUNG
   // the same network as SCL:
   #"Run Output Lamp" := "Systeem RUN";
END_REGION
END_FUNCTION

FUNCTION "SiemensEnc" : Void   // FC15, STL
TITLE = Test Siemens ENCODER
{ S7_Optimized_Access := 'FALSE' }
VERSION : 0.1
BEGIN

REGION Network 1: Presettings
         L     0;  //Delete control bits
         T     %DB1.DBD0;
         T     %DB1.DBD4;
         SET;
         S     %DB1.DBX4.0;  //Open SW gate
END_REGION

REGION Network 2: Write to the control interface
END_REGION

REGION Network 3: Read from the feedback interface
   //Read 8 bytes from the 1 Count24V
   //Configured start address of inputs
         L     "Tag_25":P;
         T     %DB1.DBD8;
         L     "Tag_26":P;
         T     %DB1.DBD12;
         R     %DB1.DBX4.0;  //Close SW gate
END_REGION
END_FUNCTION

// folder: Motion

FUNCTION_BLOCK "MC_Move"   // FB10, FBD
TITLE = MC_Move
{ S7_Optimized_Access := 'FALSE' }
VERSION : 0.1
// Block moves an Axis to an Desired Position, this block comes with the brake feature. When the axis is on position it keeps the brake for a time. You can set the time in the Brake Time field.
   VAR_INPUT
      Start : Bool;
      "Desired Position" : Real;
      "Speed (50-75%)" : Int;
      "Brake on Position" : Bool;
      Acceleration : Real;
      Deacceleration : Real;
      "Drive Ready" : Bool;
      "Drive On Position" : Bool;
      "Brake Time" : Time := T#500ms;
      "Safety OK" : Bool;
   END_VAR
   VAR_OUTPUT
      Go : Bool;
      "Desired Position Out" : Real;
      "Speed Output" : Int;
      "Acceleration Out" : Real;
      "Deacceleration Out" : Real;
      "Brake Out" : Bool;
   END_VAR
   VAR_TEMP
      SR_1 : Bool;
   END_VAR
BEGIN

REGION Network 1: Start - Go To Position + Speed